REGION Network 15
   RUNG wire#powerrail
      I_Contact( "MS050-TO" )
      Coil( "MS050-TO" )
   END_RUNG
   // the same network as SCL:
   "MS050-TO" := NOT "MS050-TO";
END_REGION

REGION Network 16
   RUNG wire#powerrail
      I_Contact( "MS051-TO" )
      Coil( "MS051-TO" )
   END_RUNG
   // the same network as SCL:
   "MS051-TO" := NOT "MS051-TO";
END_REGION

REGION Network 17
   RUNG wire#powerrail
      I_Contact( "MS052-TO" )
      Coil( "MS052-TO" )
   END_RUNG
   // the same network as SCL:
   "MS052-TO" := NOT "MS052-TO";
END_REGION

REGION Network 18
   RUNG wire#powerrail
      I_Contact( "MS053-TO" )
      Coil( "MS053-TO" )
   END_RUNG
   // the same network as SCL:
   "MS053-TO" := NOT "MS053-TO";
END_REGION

REGION Network 19: Control de Iluminación Cavaleto
   RUNG wire#powerrail
      "IluminaciónMTA"()
   END_RUNG
   // the same network as SCL:
   "IluminaciónMTA"();
END_REGION
END_FUNCTION

FUNCTION "And-Byte MTA" : Void   // FC22, LAD
{ S7_Optimized_Access := 'FALSE' }
VERSION : 0.1
BEGIN

REGION Network 1
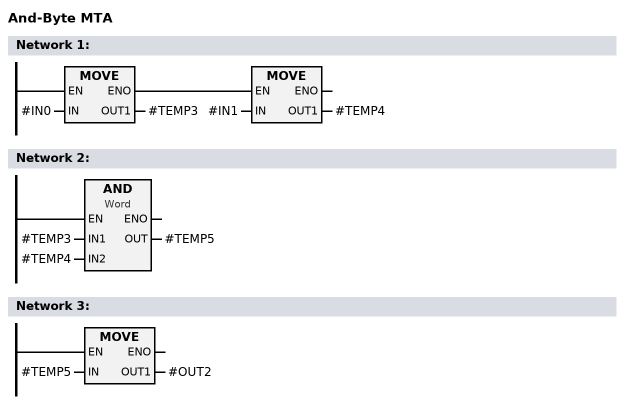
   RUNG wire#powerrail
      { S7_GenerateENO := "TRUE" } Move(in := #IN0, out1 => #TEMP3)
      { S7_GenerateENO := "TRUE" } Move(in := #IN1, out1 => #TEMP4)
   END_RUNG
   // the same network as SCL:
   // ENO of a box is taken as its EN; it also drops when the box reports an error
   #TEMP3 := #IN0;
   #TEMP4 := #IN1;
END_REGION

REGION Network 2
   RUNG wire#powerrail
      { S7_Templates := "SrcType := Word"; S7_GenerateENO := "TRUE" } And(in1 := #TEMP3, in2 := #TEMP4, out => #TEMP5)
   END_RUNG
   // the same network as SCL:
   #TEMP5 := #TEMP3 AND #TEMP4;
END_REGION

REGION Network 3
   RUNG wire#powerrail
      { S7_GenerateENO := "TRUE" } Move(in := #TEMP5, out1 => #OUT2)
   END_RUNG
   // the same network as SCL:
   #OUT2 := #TEMP5;
END_REGION
END_FUNCTION

FUNCTION "Inicialización" : Void   // FC46, LAD
{ S7_Optimized_Access := 'FALSE' }
VERSION : 0.1
BEGIN

REGION Network 1
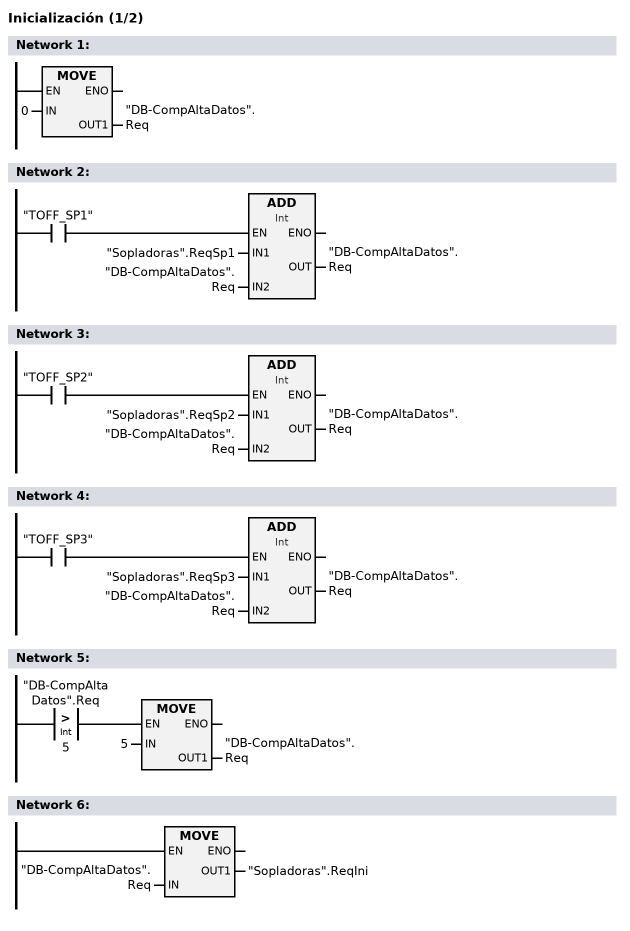
   RUNG wire#powerrail
      { S7_GenerateENO := "TRUE" } Move(in := 0, out1 => "DB-CompAltaDatos".Req)
   END_RUNG
   // the same network as SCL:
   "DB-CompAltaDatos".Req := 0;
END_REGION

REGION Network 2
   RUNG wire#powerrail
      Contact( "TOFF_SP1" )
      { S7_Templates := "SrcType := Int"; S7_GenerateENO := "TRUE" } Add(in1 := "Sopladoras".ReqSp1, in2 := "DB-CompAltaDatos".Req, out => "DB-CompAltaDatos".Req)
   END_RUNG
   // the same network as SCL:
   IF "TOFF_SP1" THEN "DB-CompAltaDatos".Req := "Sopladoras".ReqSp1 + "DB-CompAltaDatos".Req; END_IF;
END_REGION

REGION Network 3
   RUNG wire#powerrail
      Contact( "TOFF_SP2" )
      { S7_Templates := "SrcType := Int"; S7_GenerateENO := "TRUE" } Add(in1 := "Sopladoras".ReqSp2, in2 := "DB-CompAltaDatos".Req, out => "DB-CompAltaDatos".Req)
   END_RUNG
   // the same network as SCL:
   IF "TOFF_SP2" THEN "DB-CompAltaDatos".Req := "Sopladoras".ReqSp2 + "DB-CompAltaDatos".Req; END_IF;
END_REGION

REGION Network 4
   RUNG wire#powerrail
      Contact( "TOFF_SP3" )
      { S7_Templates := "SrcType := Int"; S7_GenerateENO := "TRUE" } Add(in1 := "Sopladoras".ReqSp3, in2 := "DB-CompAltaDatos".Req, out => "DB-CompAltaDatos".Req)
   END_RUNG
   // the same network as SCL:
   IF "TOFF_SP3" THEN "DB-CompAltaDatos".Req := "Sopladoras".ReqSp3 + "DB-CompAltaDatos".Req; END_IF;
END_REGION

REGION Network 5
   RUNG wire#powerrail
      { S7_Templates := "SrcType := Int" } GT_Contact(in1 := "DB-CompAltaDatos".Req, in2 := 5)
      { S7_GenerateENO := "TRUE" } Move(in := 5, out1 => "DB-CompAltaDatos".Req)
   END_RUNG
   // the same network as SCL:
   IF "DB-CompAltaDatos".Req > 5 THEN "DB-CompAltaDatos".Req := 5; END_IF;
END_REGION

REGION Network 6
   RUNG wire#powerrail
      { S7_GenerateENO := "TRUE" } Move(in := "DB-CompAltaDatos".Req, out1 => "Sopladoras".ReqIni)
   END_RUNG
   // the same network as SCL:
   "Sopladoras".ReqIni := "DB-CompAltaDatos".Req;
END_REGION

REGION Network 7
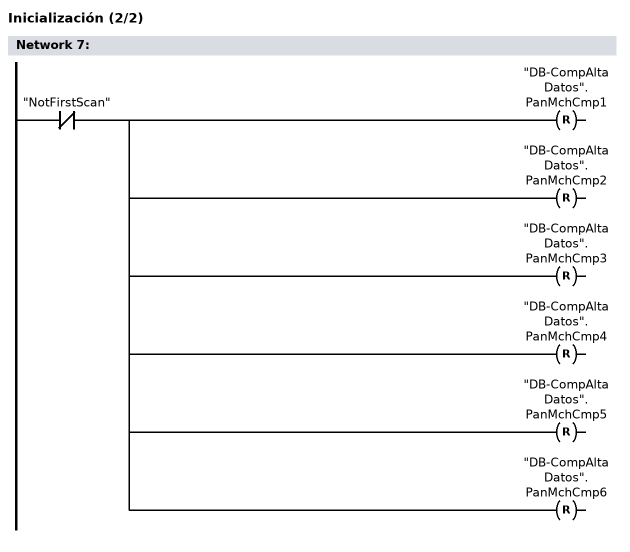
   RUNG wire#powerrail
      I_Contact( "NotFirstScan" )
      wire#w1
      R_Coil( "DB-CompAltaDatos".PanMchCmp1 )
   END_RUNG
   RUNG wire#w1
      R_Coil( "DB-CompAltaDatos".PanMchCmp2 )
   END_RUNG
   RUNG wire#w1
      R_Coil( "DB-CompAltaDatos".PanMchCmp3 )
   END_RUNG
   RUNG wire#w1
      R_Coil( "DB-CompAltaDatos".PanMchCmp4 )
   END_RUNG
   RUNG wire#w1
      R_Coil( "DB-CompAltaDatos".PanMchCmp5 )
   END_RUNG
   RUNG wire#w1
      R_Coil( "DB-CompAltaDatos".PanMchCmp6 )
   END_RUNG
   // the same network as SCL:
   IF NOT "NotFirstScan" THEN
       "DB-CompAltaDatos".PanMchCmp1 := FALSE;
       "DB-CompAltaDatos".PanMchCmp2 := FALSE;
       "DB-CompAltaDatos".PanMchCmp3 := FALSE;
       "DB-CompAltaDatos".PanMchCmp4 := FALSE;
       "DB-CompAltaDatos".PanMchCmp5 := FALSE;
       "DB-CompAltaDatos".PanMchCmp6 := FALSE;
   END_IF;
END_REGION
END_FUNCTION

// folder: Bloques Estándar

FUNCTION_BLOCK "ControladorMotoresMTA"   // FB2, LAD
{ S7_Optimized_Access := 'FALSE' }
VERSION : 0.1
BEGIN

REGION Network 2
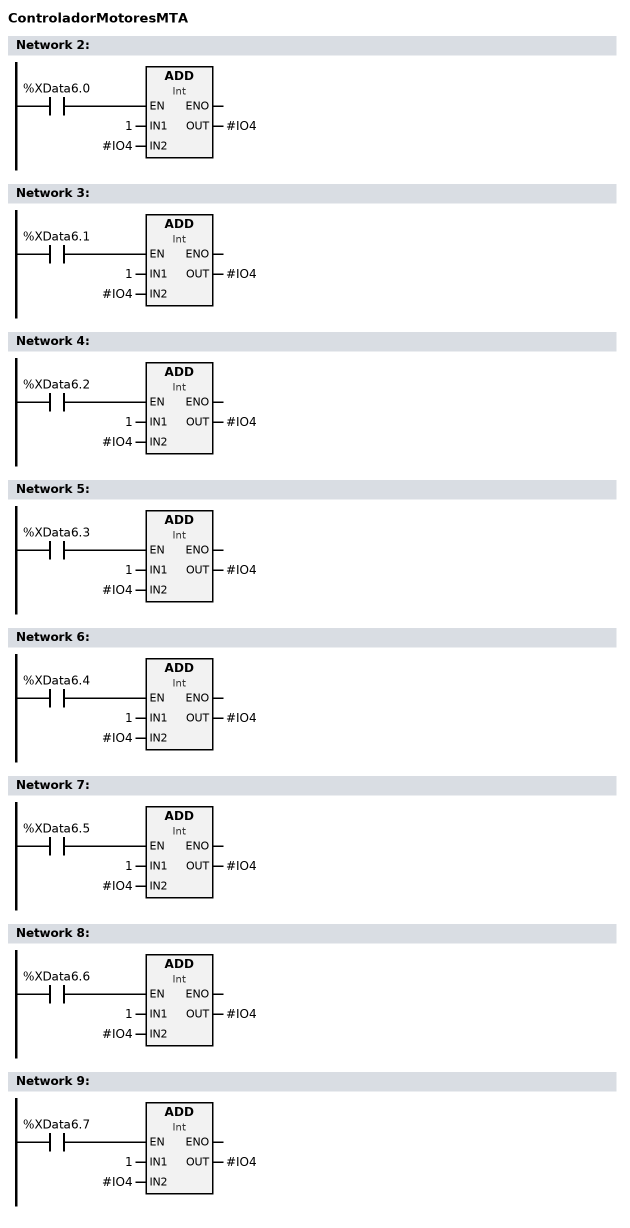
   RUNG wire#powerrail
      Contact( %XData6.0 )
      { S7_Templates := "SrcType := Int"; S7_GenerateENO := "TRUE" } Add(in1 := 1, in2 := #IO4, out => #IO4)
   END_RUNG
   // the same network as SCL:
   IF %XData6.0 THEN #IO4 := 1 + #IO4; END_IF;
END_REGION

REGION Network 3
   RUNG wire#powerrail
      Contact( %XData6.1 )
      { S7_Templates := "SrcType := Int"; S7_GenerateENO := "TRUE" } Add(in1 := 1, in2 := #IO4, out => #IO4)
   END_RUNG
   // the same network as SCL:
   IF %XData6.1 THEN #IO4 := 1 + #IO4; END_IF;
END_REGION

REGION Network 4
   RUNG wire#powerrail
      Contact( %XData6.2 )
      { S7_Templates := "SrcType := Int"; S7_GenerateENO := "TRUE" } Add(in1 := 1, in2 := #IO4, out => #IO4)
   END_RUNG
   // the same network as SCL:
   IF %XData6.2 THEN #IO4 := 1 + #IO4; END_IF;
END_REGION

REGION Network 5
   RUNG wire#powerrail
      Contact( %XData6.3 )
      { S7_Templates := "SrcType := Int"; S7_GenerateENO := "TRUE" } Add(in1 := 1, in2 := #IO4, out => #IO4)
   END_RUNG
   // the same network as SCL:
   IF %XData6.3 THEN #IO4 := 1 + #IO4; END_IF;
END_REGION

REGION Network 6
   RUNG wire#powerrail
      Contact( %XData6.4 )
      { S7_Templates := "SrcType := Int"; S7_GenerateENO := "TRUE" } Add(in1 := 1, in2 := #IO4, out => #IO4)
   END_RUNG
   // the same network as SCL:
   IF %XData6.4 THEN #IO4 := 1 + #IO4; END_IF;
END_REGION

REGION Network 7
   RUNG wire#powerrail
      Contact( %XData6.5 )
      { S7_Templates := "SrcType := Int"; S7_GenerateENO := "TRUE" } Add(in1 := 1, in2 := #IO4, out => #IO4)
   END_RUNG
   // the same network as SCL:
   IF %XData6.5 THEN #IO4 := 1 + #IO4; END_IF;
END_REGION

REGION Network 8
   RUNG wire#powerrail
      Contact( %XData6.6 )
      { S7_Templates := "SrcType := Int"; S7_GenerateENO := "TRUE" } Add(in1 := 1, in2 := #IO4, out => #IO4)
   END_RUNG
   // the same network as SCL:
   IF %XData6.6 THEN #IO4 := 1 + #IO4; END_IF;
END_REGION

REGION Network 9
   RUNG wire#powerrail
      Contact( %XData6.7 )
      { S7_Templates := "SrcType := Int"; S7_GenerateENO := "TRUE" } Add(in1 := 1, in2 := #IO4, out => #IO4)
   END_RUNG
   // the same network as SCL:
   IF %XData6.7 THEN #IO4 := 1 + #IO4; END_IF;
END_REGION
END_FUNCTION_BLOCK

// folder: Bloques Estándar/Boosters

FUNCTION "Booster (MTA)" : Void   // FC25, LAD
TITLE = Manejo General de los Boosters
{ S7_Optimized_Access := 'FALSE' }
VERSION : 0.1
   VAR_TEMP   // added for the SCL form of the ladder/FBD networks
      _w1 : Bool;
      _s5time1 : S5Time;
      _w2 : Bool;
      _s5time2 : S5Time;
      _w3 : Bool;
   END_VAR
BEGIN

REGION Network 1: Validación Horas para invertir prioridades
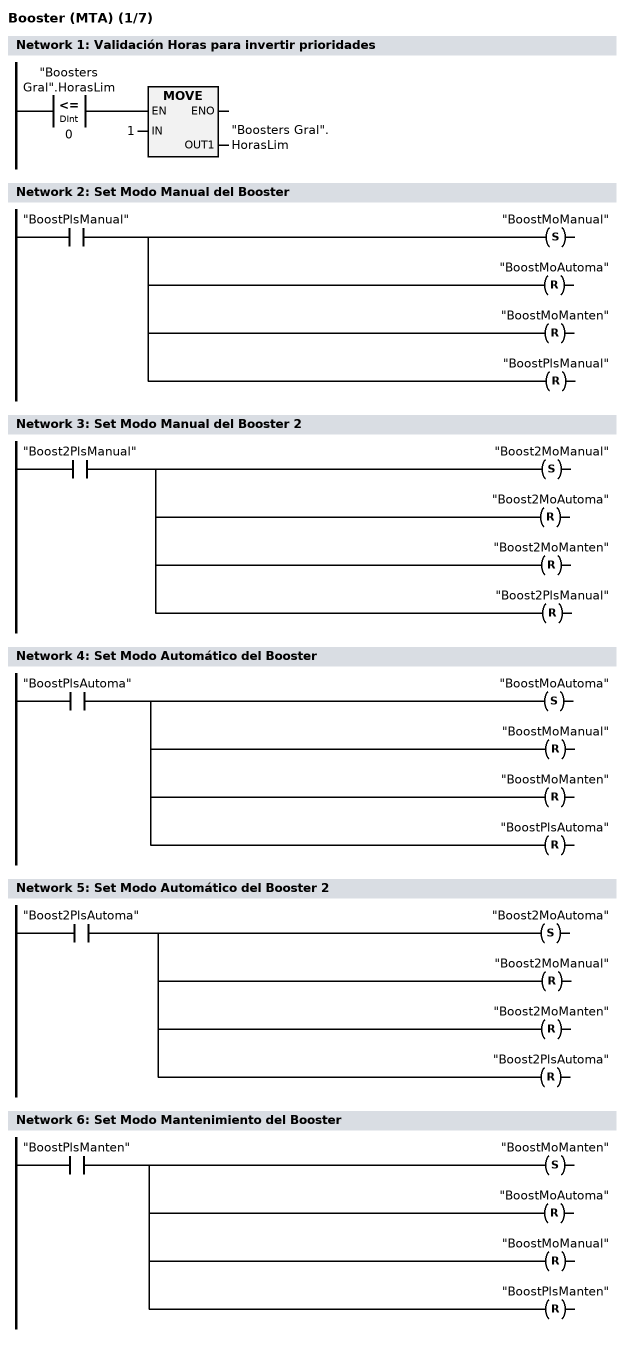
   RUNG wire#powerrail
      { S7_Templates := "SrcType := DInt" } LE_Contact(in1 := "Boosters Gral".HorasLim, in2 := 0)
      { S7_GenerateENO := "TRUE" } Move(in := 1, out1 => "Boosters Gral".HorasLim)
   END_RUNG
   // the same network as SCL:
   IF "Boosters Gral".HorasLim <= 0 THEN "Boosters Gral".HorasLim := 1; END_IF;
END_REGION

REGION Network 2: Set Modo Manual del Booster
   RUNG wire#powerrail
      Contact( "BoostPlsManual" )
      wire#w1
      S_Coil( "BoostMoManual" )
   END_RUNG
   RUNG wire#w1
      R_Coil( "BoostMoAutoma" )
   END_RUNG
   RUNG wire#w1
      R_Coil( "BoostMoManten" )
   END_RUNG
   RUNG wire#w1
      R_Coil( "BoostPlsManual" )
   END_RUNG
   // the same network as SCL:
   IF "BoostPlsManual" THEN
       "BoostMoManual" := TRUE;
       "BoostMoAutoma" := FALSE;
       "BoostMoManten" := FALSE;
       "BoostPlsManual" := FALSE;
   END_IF;
END_REGION

REGION Network 3: Set Modo Manual del Booster 2
   RUNG wire#powerrail
      Contact( "Boost2PlsManual" )
      wire#w1
      S_Coil( "Boost2MoManual" )
   END_RUNG
   RUNG wire#w1
      R_Coil( "Boost2MoAutoma" )
   END_RUNG
   RUNG wire#w1
      R_Coil( "Boost2MoManten" )
   END_RUNG
   RUNG wire#w1
      R_Coil( "Boost2PlsManual" )
   END_RUNG
   // the same network as SCL:
   IF "Boost2PlsManual" THEN
       "Boost2MoManual" := TRUE;
       "Boost2MoAutoma" := FALSE;
       "Boost2MoManten" := FALSE;
       "Boost2PlsManual" := FALSE;
   END_IF;
END_REGION

REGION Network 4: Set Modo Automático del Booster
   RUNG wire#powerrail
      Contact( "BoostPlsAutoma" )
      wire#w1
      S_Coil( "BoostMoAutoma" )
   END_RUNG
   RUNG wire#w1
      R_Coil( "BoostMoManual" )
   END_RUNG
   RUNG wire#w1
      R_Coil( "BoostMoManten" )
   END_RUNG
   RUNG wire#w1
      R_Coil( "BoostPlsAutoma" )
   END_RUNG
   // the same network as SCL:
   IF "BoostPlsAutoma" THEN
       "BoostMoAutoma" := TRUE;
       "BoostMoManual" := FALSE;
       "BoostMoManten" := FALSE;
       "BoostPlsAutoma" := FALSE;
   END_IF;
END_REGION

REGION Network 5: Set Modo Automático del Booster 2
   RUNG wire#powerrail
      Contact( "Boost2PlsAutoma" )
      wire#w1
      S_Coil( "Boost2MoAutoma" )
   END_RUNG
   RUNG wire#w1
      R_Coil( "Boost2MoManual" )
   END_RUNG
   RUNG wire#w1
      R_Coil( "Boost2MoManten" )
   END_RUNG
   RUNG wire#w1
      R_Coil( "Boost2PlsAutoma" )
   END_RUNG
   // the same network as SCL:
   IF "Boost2PlsAutoma" THEN
       "Boost2MoAutoma" := TRUE;
       "Boost2MoManual" := FALSE;
       "Boost2MoManten" := FALSE;
       "Boost2PlsAutoma" := FALSE;
   END_IF;
END_REGION

REGION Network 6: Set Modo Mantenimiento del Booster
   RUNG wire#powerrail
      Contact( "BoostPlsManten" )
      wire#w1
      S_Coil( "BoostMoManten" )
   END_RUNG
   RUNG wire#w1
      R_Coil( "BoostMoAutoma" )
   END_RUNG
   RUNG wire#w1
      R_Coil( "BoostMoManual" )
   END_RUNG
   RUNG wire#w1
      R_Coil( "BoostPlsManten" )
   END_RUNG
   // the same network as SCL:
   IF "BoostPlsManten" THEN
       "BoostMoManten" := TRUE;
       "BoostMoAutoma" := FALSE;
       "BoostMoManual" := FALSE;
       "BoostPlsManten" := FALSE;
   END_IF;
END_REGION

REGION Network 7: Set Modo Mantenimiento del Booster 2
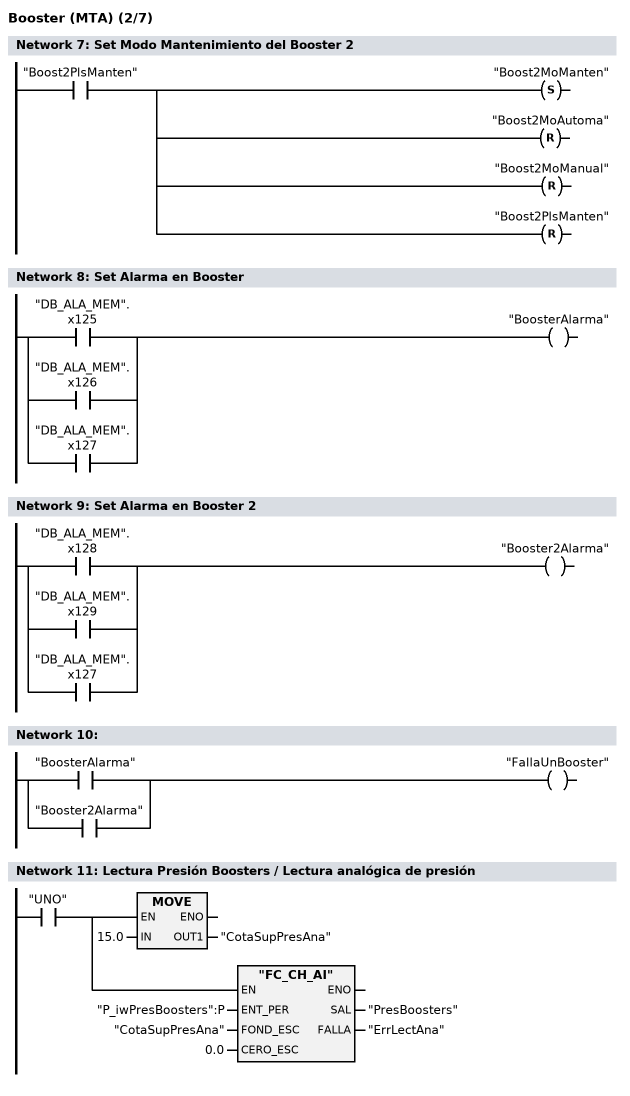
   RUNG wire#powerrail
      Contact( "Boost2PlsManten" )
      wire#w1
      S_Coil( "Boost2MoManten" )
   END_RUNG
   RUNG wire#w1
      R_Coil( "Boost2MoAutoma" )
   END_RUNG
   RUNG wire#w1
      R_Coil( "Boost2MoManual" )
   END_RUNG
   RUNG wire#w1
      R_Coil( "Boost2PlsManten" )
   END_RUNG
   // the same network as SCL:
   IF "Boost2PlsManten" THEN
       "Boost2MoManten" := TRUE;
       "Boost2MoAutoma" := FALSE;
       "Boost2MoManual" := FALSE;
       "Boost2PlsManten" := FALSE;
   END_IF;
END_REGION

REGION Network 8: Set Alarma en Booster
   RUNG wire#powerrail
      Contact( "DB_ALA_MEM".x125 )
      wire#w1
      Coil( "BoosterAlarma" )
   END_RUNG
   RUNG wire#powerrail
      Contact( "DB_ALA_MEM".x126 )
   END_RUNG wire#w1
   RUNG wire#powerrail
      Contact( "DB_ALA_MEM".x127 )
   END_RUNG wire#w1
   // the same network as SCL:
   "BoosterAlarma" := "DB_ALA_MEM".x125 OR "DB_ALA_MEM".x126 OR "DB_ALA_MEM".x127;
END_REGION

REGION Network 9: Set Alarma en Booster 2
   RUNG wire#powerrail
      Contact( "DB_ALA_MEM".x128 )
      wire#w1
      Coil( "Booster2Alarma" )
   END_RUNG
   RUNG wire#powerrail
      Contact( "DB_ALA_MEM".x129 )
   END_RUNG wire#w1
   RUNG wire#powerrail
      Contact( "DB_ALA_MEM".x127 )
   END_RUNG wire#w1
   // the same network as SCL:
   "Booster2Alarma" := "DB_ALA_MEM".x128 OR "DB_ALA_MEM".x129 OR "DB_ALA_MEM".x127;
END_REGION

REGION Network 10
   RUNG wire#powerrail
      Contact( "BoosterAlarma" )
      wire#w1
      Coil( "FallaUnBooster" )
   END_RUNG
   RUNG wire#powerrail
      Contact( "Booster2Alarma" )
   END_RUNG wire#w1
   // the same network as SCL:
   "FallaUnBooster" := "BoosterAlarma" OR "Booster2Alarma";
END_REGION

REGION Network 11: Lectura Presión Boosters / Lectura analógica de presión
   RUNG wire#powerrail
      Contact( "UNO" )
      wire#w1
      { S7_GenerateENO := "TRUE" } Move(in := 15.0, out1 => "CotaSupPresAna")
   END_RUNG
   RUNG wire#w1
      "FC_CH_AI"(ENT_PER := "P_iwPresBoosters":P, FOND_ESC := "CotaSupPresAna", CERO_ESC := 0.0, SAL => "PresBoosters", FALLA => "ErrLectAna")
   END_RUNG
   // the same network as SCL:
   IF "UNO" THEN
       "CotaSupPresAna" := 15.0;
       "FC_CH_AI"(ENT_PER := "P_iwPresBoosters":P,
                  FOND_ESC := "CotaSupPresAna",
                  CERO_ESC := 0.0,
                  SAL => "PresBoosters",
                  FALLA => "ErrLectAna");
   END_IF;
END_REGION

REGION Network 12: Bandas de presión para arranque de Boosters / Set-Reset para control analógico
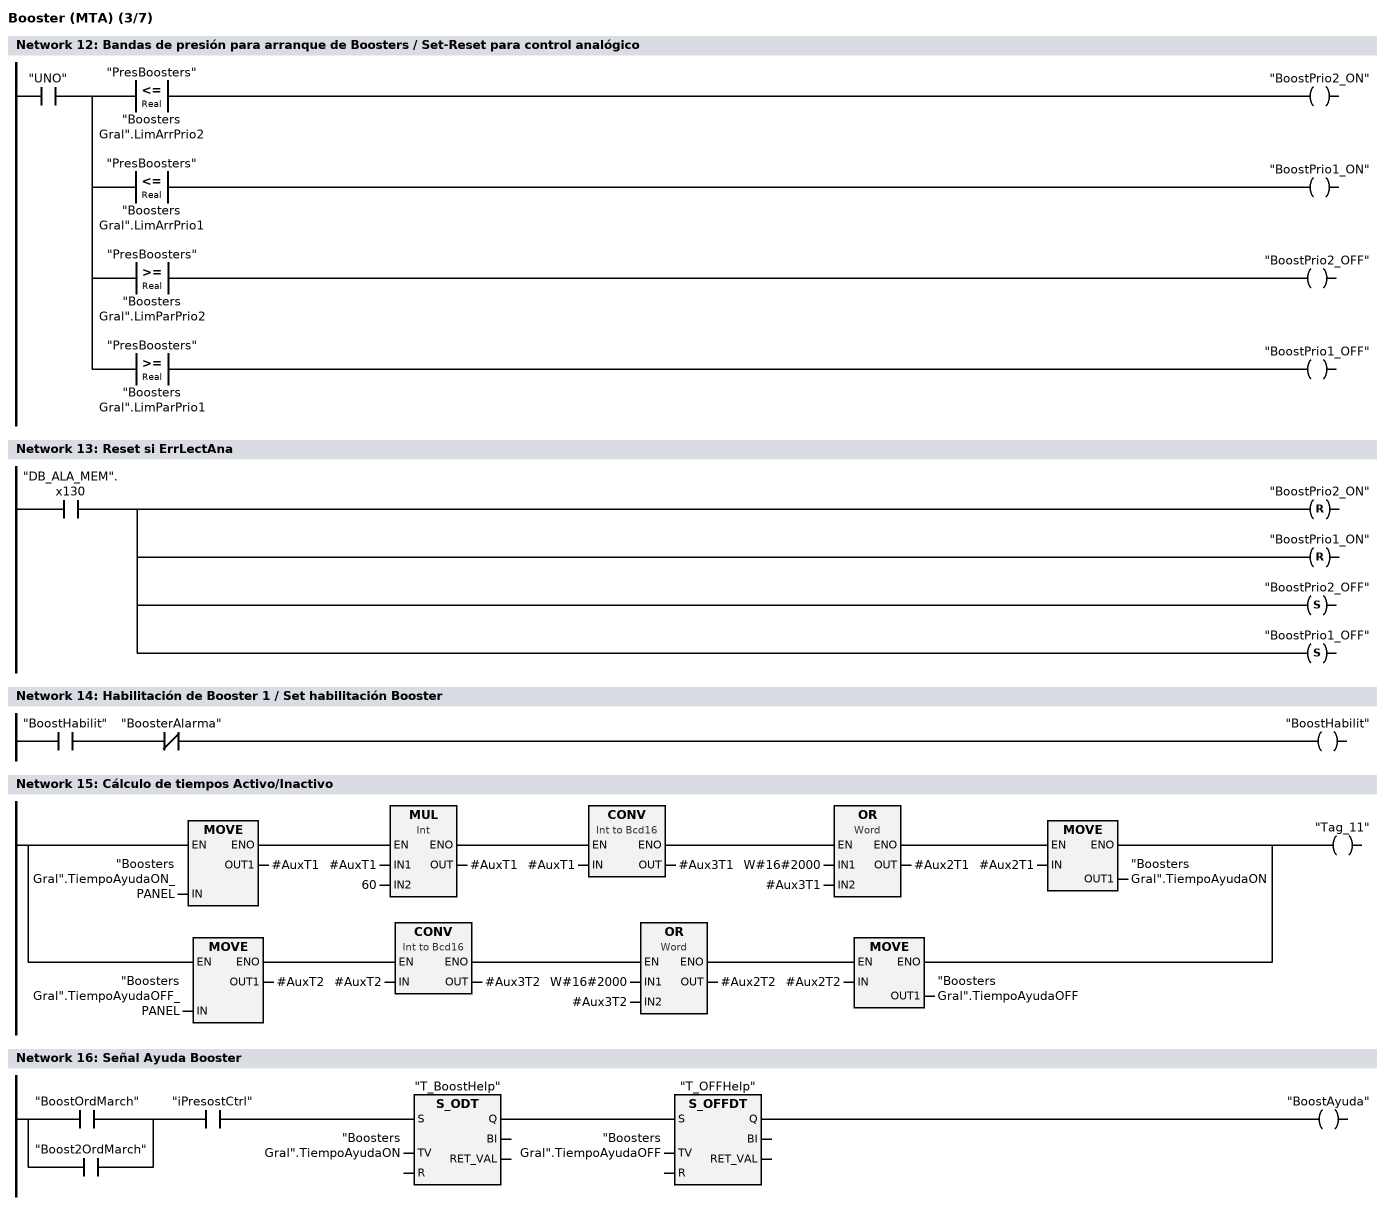
   RUNG wire#powerrail
      Contact( "UNO" )
      wire#w1
      { S7_Templates := "SrcType := Real" } LE_Contact(in1 := "PresBoosters", in2 := "Boosters Gral".LimArrPrio2)
      Coil( "BoostPrio2_ON" )
   END_RUNG
   RUNG wire#w1
      { S7_Templates := "SrcType := Real" } LE_Contact(in1 := "PresBoosters", in2 := "Boosters Gral".LimArrPrio1)
      Coil( "BoostPrio1_ON" )
   END_RUNG
   RUNG wire#w1
      { S7_Templates := "SrcType := Real" } GE_Contact(in1 := "PresBoosters", in2 := "Boosters Gral".LimParPrio2)
      Coil( "BoostPrio2_OFF" )
   END_RUNG
   RUNG wire#w1
      { S7_Templates := "SrcType := Real" } GE_Contact(in1 := "PresBoosters", in2 := "Boosters Gral".LimParPrio1)
      Coil( "BoostPrio1_OFF" )
   END_RUNG
   // the same network as SCL:
   "BoostPrio2_ON" := "UNO" AND ("PresBoosters" <= "Boosters Gral".LimArrPrio2);
   "BoostPrio1_ON" := "UNO" AND ("PresBoosters" <= "Boosters Gral".LimArrPrio1);
   "BoostPrio2_OFF" := "UNO" AND ("PresBoosters" >= "Boosters Gral".LimParPrio2);
   "BoostPrio1_OFF" := "UNO" AND ("PresBoosters" >= "Boosters Gral".LimParPrio1);
END_REGION

REGION Network 13: Reset si ErrLectAna
   RUNG wire#powerrail
      Contact( "DB_ALA_MEM".x130 )
      wire#w1
      R_Coil( "BoostPrio2_ON" )
   END_RUNG
   RUNG wire#w1
      R_Coil( "BoostPrio1_ON" )
   END_RUNG
   RUNG wire#w1
      S_Coil( "BoostPrio2_OFF" )
   END_RUNG
   RUNG wire#w1
      S_Coil( "BoostPrio1_OFF" )
   END_RUNG
   // the same network as SCL:
   IF "DB_ALA_MEM".x130 THEN
       "BoostPrio2_ON" := FALSE;
       "BoostPrio1_ON" := FALSE;
       "BoostPrio2_OFF" := TRUE;
       "BoostPrio1_OFF" := TRUE;
   END_IF;
END_REGION

REGION Network 14: Habilitación de Booster 1 / Set habilitación Booster
   RUNG wire#powerrail
      Contact( "BoostHabilit" )
      I_Contact( "BoosterAlarma" )
      Coil( "BoostHabilit" )
   END_RUNG
   // the same network as SCL:
   "BoostHabilit" := "BoostHabilit" AND NOT "BoosterAlarma";
END_REGION

REGION Network 15: Cálculo de tiempos Activo/Inactivo
   // no checked SCL form for this network; see the picture
END_REGION

REGION Network 16: Señal Ayuda Booster
   RUNG wire#powerrail
      Contact( "BoostOrdMarch" )
      wire#w1
      Contact( "iPresostCtrl" )
      S_ODT(T_NO := "T_BoostHelp", TV := "Boosters Gral".TiempoAyudaON, R :=, BI =>, RET_VAL =>)
      S_OFFDT(T_NO := "T_OFFHelp", TV := "Boosters Gral".TiempoAyudaOFF, R :=, BI =>, RET_VAL =>)
      Coil( "BoostAyuda" )
   END_RUNG
   RUNG wire#powerrail
      Contact( "Boost2OrdMarch" )
   END_RUNG wire#w1
   // the same network as SCL:
   #_s5time1 := S_ODT(T_NO := "T_BoostHelp",
                      S := ("BoostOrdMarch" OR "Boost2OrdMarch") AND "iPresostCtrl",
                      TV := "Boosters Gral".TiempoAyudaON,
                      Q => #_w1);
   #_s5time2 := S_OFFDT(T_NO := "T_OFFHelp", S := #_w1, TV := "Boosters Gral".TiempoAyudaOFF, Q => #_w2);
   "BoostAyuda" := #_w2;
END_REGION

REGION Network 17: Prioridades Boosters / Prioridades Nulas
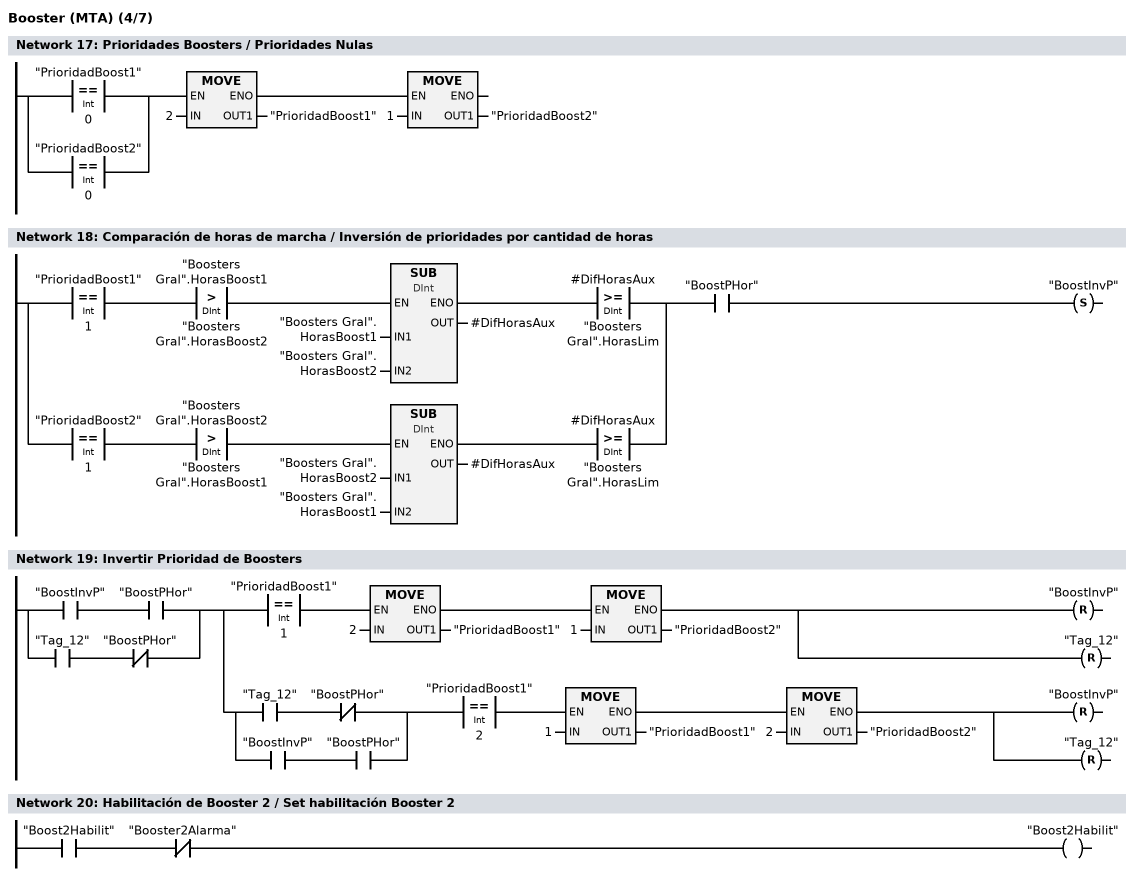
   RUNG wire#powerrail
      { S7_Templates := "SrcType := Int" } EQ_Contact(in1 := "PrioridadBoost1", in2 := 0)
      wire#w1
      { S7_GenerateENO := "TRUE" } Move(in := 2, out1 => "PrioridadBoost1")
      { S7_GenerateENO := "TRUE" } Move(in := 1, out1 => "PrioridadBoost2")
   END_RUNG
   RUNG wire#powerrail
      { S7_Templates := "SrcType := Int" } EQ_Contact(in1 := "PrioridadBoost2", in2 := 0)
   END_RUNG wire#w1
   // the same network as SCL:
   // ENO of a box is taken as its EN; it also drops when the box reports an error
   #_w1 := ("PrioridadBoost1" = 0) OR ("PrioridadBoost2" = 0);
   IF #_w1 THEN
       "PrioridadBoost1" := 2;
       "PrioridadBoost2" := 1;
   END_IF;
END_REGION

REGION Network 18: Comparación de horas de marcha / Inversión de prioridades por cantidad de horas
   RUNG wire#powerrail
      { S7_Templates := "SrcType := Int" } EQ_Contact(in1 := "PrioridadBoost1", in2 := 1)
      { S7_Templates := "SrcType := DInt" } GT_Contact(in1 := "Boosters Gral".HorasBoost1, in2 := "Boosters Gral".HorasBoost2)
      { S7_Templates := "SrcType := DInt"; S7_GenerateENO := "TRUE" } Sub(in1 := "Boosters Gral".HorasBoost1, in2 := "Boosters Gral".HorasBoost2, out => #DifHorasAux)
      { S7_Templates := "SrcType := DInt" } GE_Contact(in1 := #DifHorasAux, in2 := "Boosters Gral".HorasLim)
      wire#w1
      Contact( "BoostPHor" )
      S_Coil( "BoostInvP" )
   END_RUNG
   RUNG wire#powerrail
      { S7_Templates := "SrcType := Int" } EQ_Contact(in1 := "PrioridadBoost2", in2 := 1)
      { S7_Templates := "SrcType := DInt" } GT_Contact(in1 := "Boosters Gral".HorasBoost2, in2 := "Boosters Gral".HorasBoost1)
      { S7_Templates := "SrcType := DInt"; S7_GenerateENO := "TRUE" } Sub(in1 := "Boosters Gral".HorasBoost2, in2 := "Boosters Gral".HorasBoost1, out => #DifHorasAux)
      { S7_Templates := "SrcType := DInt" } GE_Contact(in1 := #DifHorasAux, in2 := "Boosters Gral".HorasLim)
   END_RUNG wire#w1
   // the same network as SCL:
   // ENO of a box is taken as its EN; it also drops when the box reports an error
   #_w1 := ("PrioridadBoost1" = 1) AND ("Boosters Gral".HorasBoost1 > "Boosters Gral".HorasBoost2);
   IF #_w1 THEN #DifHorasAux := "Boosters Gral".HorasBoost1 - "Boosters Gral".HorasBoost2; END_IF;
   #_w2 := ("PrioridadBoost2" = 1) AND ("Boosters Gral".HorasBoost2 > "Boosters Gral".HorasBoost1);
   #_w3 := #_w1 AND (#DifHorasAux >= "Boosters Gral".HorasLim);
   IF #_w2 THEN #DifHorasAux := "Boosters Gral".HorasBoost2 - "Boosters Gral".HorasBoost1; END_IF;
   IF (#_w3 OR (#_w2 AND (#DifHorasAux >= "Boosters Gral".HorasLim))) AND "BoostPHor" THEN
       "BoostInvP" := TRUE;
   END_IF;
END_REGION

REGION Network 19: Invertir Prioridad de Boosters
   RUNG wire#powerrail
      Contact( "BoostInvP" )
      Contact( "BoostPHor" )
      wire#w1
      { S7_Templates := "SrcType := Int" } EQ_Contact(in1 := "PrioridadBoost1", in2 := 1)
      { S7_GenerateENO := "TRUE" } Move(in := 2, out1 => "PrioridadBoost1")
      { S7_GenerateENO := "TRUE" } Move(in := 1, out1 => "PrioridadBoost2")
      wire#w2
      R_Coil( "BoostInvP" )
   END_RUNG
   RUNG wire#powerrail
      Contact( "Tag_12" )
      I_Contact( "BoostPHor" )
   END_RUNG wire#w1
   RUNG wire#w2
      R_Coil( "Tag_12" )
   END_RUNG
   RUNG wire#w1
      Contact( "Tag_12" )
      I_Contact( "BoostPHor" )
      wire#w3
      { S7_Templates := "SrcType := Int" } EQ_Contact(in1 := "PrioridadBoost1", in2 := 2)
      { S7_GenerateENO := "TRUE" } Move(in := 1, out1 => "PrioridadBoost1")
      { S7_GenerateENO := "TRUE" } Move(in := 2, out1 => "PrioridadBoost2")
      wire#w4
      R_Coil( "BoostInvP" )
   END_RUNG
   RUNG wire#w1
      Contact( "BoostInvP" )
      Contact( "BoostPHor" )
   END_RUNG wire#w3
   RUNG wire#w4
      R_Coil( "Tag_12" )
   END_RUNG
   // the same network as SCL:
   // ENO of a box is taken as its EN; it also drops when the box reports an error
   #_w1 := ("BoostInvP" AND "BoostPHor") OR ("Tag_12" AND NOT "BoostPHor");
   #_w2 := #_w1 AND ("PrioridadBoost1" = 1);
   IF #_w2 THEN
       "PrioridadBoost1" := 2;
       "PrioridadBoost2" := 1;
       "BoostInvP" := FALSE;
       "Tag_12" := FALSE;
   END_IF;
   #_w3 := #_w1 AND (("Tag_12" AND NOT "BoostPHor") OR ("BoostInvP" AND "BoostPHor")) AND ("PrioridadBoost1" = 2);
   IF #_w3 THEN
       "PrioridadBoost1" := 1;
       "PrioridadBoost2" := 2;
       "BoostInvP" := FALSE;
       "Tag_12" := FALSE;
   END_IF;
END_REGION

REGION Network 20: Habilitación de Booster 2 / Set habilitación Booster 2
   RUNG wire#powerrail
      Contact( "Boost2Habilit" )
      I_Contact( "Booster2Alarma" )
      Coil( "Boost2Habilit" )
   END_RUNG
   // the same network as SCL:
   "Boost2Habilit" := "Boost2Habilit" AND NOT "Booster2Alarma";
END_REGION

REGION Network 21: Orden de Marcha Booster
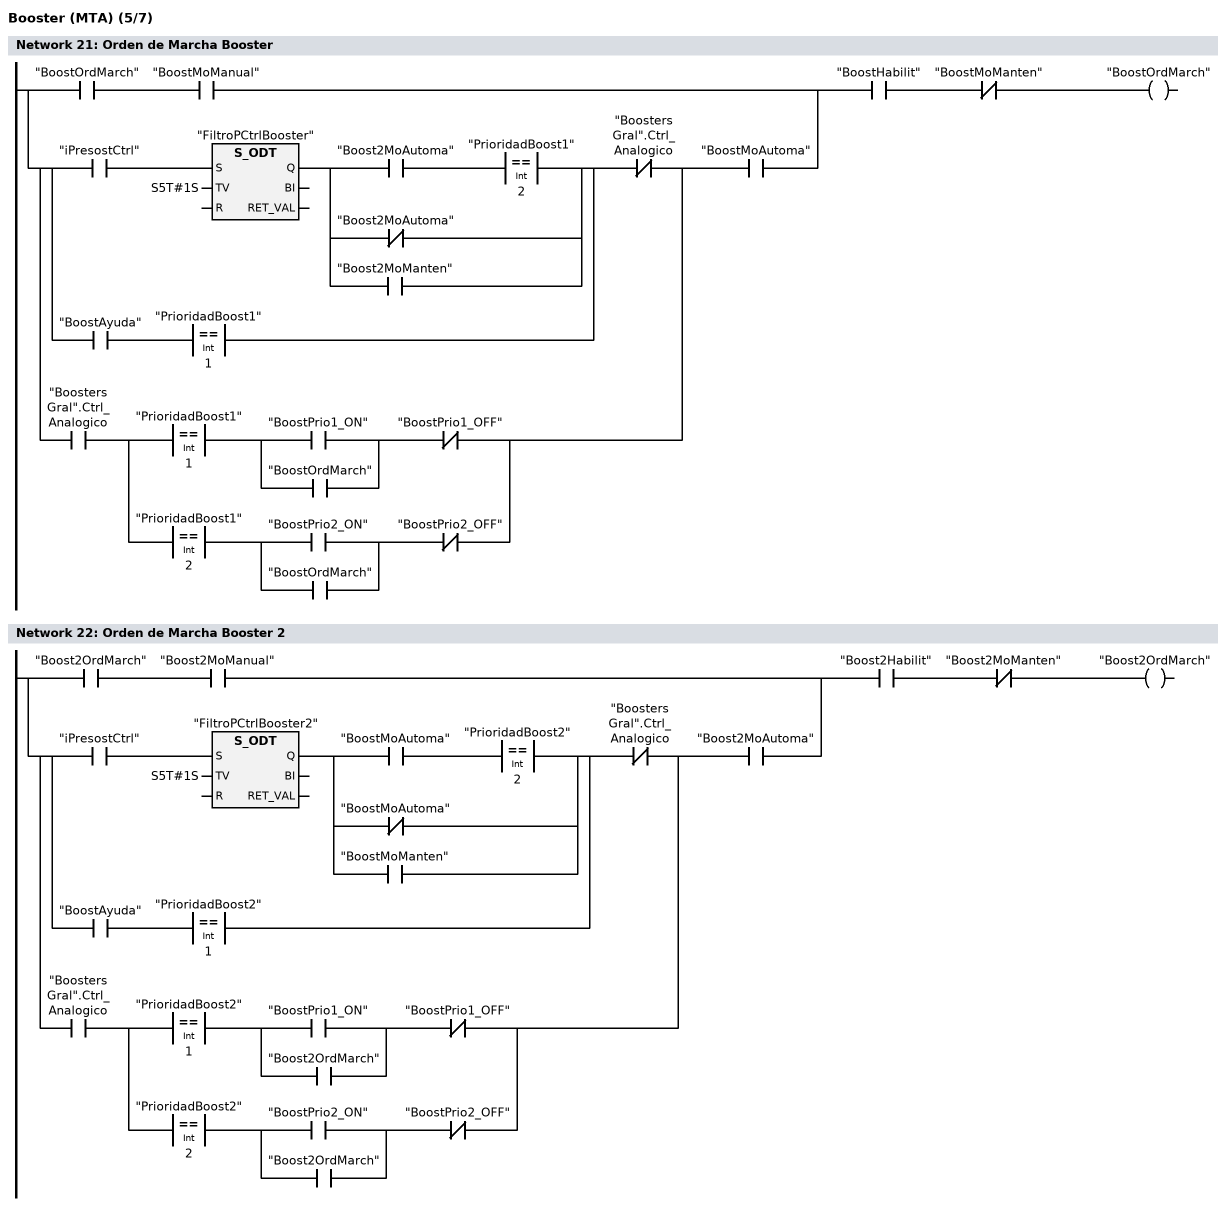
   RUNG wire#powerrail
      Contact( "BoostOrdMarch" )
      Contact( "BoostMoManual" )
      wire#w1
      Contact( "BoostHabilit" )
      I_Contact( "BoostMoManten" )
      Coil( "BoostOrdMarch" )
   END_RUNG
   RUNG wire#powerrail
      Contact( "iPresostCtrl" )
      S_ODT(T_NO := "FiltroPCtrlBooster", TV := S5T#1S, R :=, BI =>, RET_VAL =>)
      wire#w2
      Contact( "Boost2MoAutoma" )
      { S7_Templates := "SrcType := Int" } EQ_Contact(in1 := "PrioridadBoost1", in2 := 2)
      wire#w3
      I_Contact( "Boosters Gral".Ctrl_Analogico )
      wire#w4
      Contact( "BoostMoAutoma" )
   END_RUNG wire#w1
   RUNG wire#w2
      I_Contact( "Boost2MoAutoma" )
   END_RUNG wire#w3
   RUNG wire#w2
      Contact( "Boost2MoManten" )
   END_RUNG wire#w3
   RUNG wire#powerrail
      Contact( "BoostAyuda" )
      { S7_Templates := "SrcType := Int" } EQ_Contact(in1 := "PrioridadBoost1", in2 := 1)
   END_RUNG wire#w3
   RUNG wire#powerrail
      Contact( "Boosters Gral".Ctrl_Analogico )
      wire#w5
      { S7_Templates := "SrcType := Int" } EQ_Contact(in1 := "PrioridadBoost1", in2 := 1)
      wire#w6
      Contact( "BoostPrio1_ON" )
      wire#w7
      I_Contact( "BoostPrio1_OFF" )
   END_RUNG wire#w4
   RUNG wire#w6
      Contact( "BoostOrdMarch" )
   END_RUNG wire#w7
   RUNG wire#w5
      { S7_Templates := "SrcType := Int" } EQ_Contact(in1 := "PrioridadBoost1", in2 := 2)
      wire#w8
      Contact( "BoostPrio2_ON" )
      wire#w9
      I_Contact( "BoostPrio2_OFF" )
   END_RUNG wire#w4
   RUNG wire#w8
      Contact( "BoostOrdMarch" )
   END_RUNG wire#w9
   // the same network as SCL:
   #_s5time1 := S_ODT(T_NO := "FiltroPCtrlBooster", S := "iPresostCtrl", TV := S5T#1S, Q => #_w1);
   "BoostOrdMarch" := (("BoostOrdMarch" AND "BoostMoManual") OR (((((#_w1 AND (("Boost2MoAutoma" AND ("PrioridadBoost1" = 2)) OR NOT "Boost2MoAutoma" OR "Boost2MoManten")) OR ("BoostAyuda" AND ("PrioridadBoost1" = 1))) AND NOT "Boosters Gral".Ctrl_Analogico) OR ("Boosters Gral".Ctrl_Analogico AND ((("PrioridadBoost1" = 1) AND ("BoostPrio1_ON" OR "BoostOrdMarch") AND NOT "BoostPrio1_OFF") OR (("PrioridadBoost1" = 2) AND ("BoostPrio2_ON" OR "BoostOrdMarch") AND NOT "BoostPrio2_OFF")))) AND "BoostMoAutoma")) AND "BoostHabilit" AND NOT "BoostMoManten";
END_REGION

REGION Network 22: Orden de Marcha Booster 2
   RUNG wire#powerrail
      Contact( "Boost2OrdMarch" )
      Contact( "Boost2MoManual" )
      wire#w1
      Contact( "Boost2Habilit" )
      I_Contact( "Boost2MoManten" )
      Coil( "Boost2OrdMarch" )
   END_RUNG
   RUNG wire#powerrail
      Contact( "iPresostCtrl" )
      S_ODT(T_NO := "FiltroPCtrlBooster2", TV := S5T#1S, R :=, BI =>, RET_VAL =>)
      wire#w2
      Contact( "BoostMoAutoma" )
      { S7_Templates := "SrcType := Int" } EQ_Contact(in1 := "PrioridadBoost2", in2 := 2)
      wire#w3
      I_Contact( "Boosters Gral".Ctrl_Analogico )
      wire#w4
      Contact( "Boost2MoAutoma" )
   END_RUNG wire#w1
   RUNG wire#w2
      I_Contact( "BoostMoAutoma" )
   END_RUNG wire#w3
   RUNG wire#w2
      Contact( "BoostMoManten" )
   END_RUNG wire#w3
   RUNG wire#powerrail
      Contact( "BoostAyuda" )
      { S7_Templates := "SrcType := Int" } EQ_Contact(in1 := "PrioridadBoost2", in2 := 1)
   END_RUNG wire#w3
   RUNG wire#powerrail
      Contact( "Boosters Gral".Ctrl_Analogico )
      wire#w5
      { S7_Templates := "SrcType := Int" } EQ_Contact(in1 := "PrioridadBoost2", in2 := 1)
      wire#w6
      Contact( "BoostPrio1_ON" )
      wire#w7
      I_Contact( "BoostPrio1_OFF" )
   END_RUNG wire#w4
   RUNG wire#w6
      Contact( "Boost2OrdMarch" )
   END_RUNG wire#w7
   RUNG wire#w5
      { S7_Templates := "SrcType := Int" } EQ_Contact(in1 := "PrioridadBoost2", in2 := 2)
      wire#w8
      Contact( "BoostPrio2_ON" )
      wire#w9
      I_Contact( "BoostPrio2_OFF" )
   END_RUNG wire#w4
   RUNG wire#w8
      Contact( "Boost2OrdMarch" )
   END_RUNG wire#w9
   // the same network as SCL:
   #_s5time1 := S_ODT(T_NO := "FiltroPCtrlBooster2", S := "iPresostCtrl", TV := S5T#1S, Q => #_w1);
   "Boost2OrdMarch" := (("Boost2OrdMarch" AND "Boost2MoManual") OR (((((#_w1 AND (("BoostMoAutoma" AND ("PrioridadBoost2" = 2)) OR NOT "BoostMoAutoma" OR "BoostMoManten")) OR ("BoostAyuda" AND ("PrioridadBoost2" = 1))) AND NOT "Boosters Gral".Ctrl_Analogico) OR ("Boosters Gral".Ctrl_Analogico AND ((("PrioridadBoost2" = 1) AND ("BoostPrio1_ON" OR "Boost2OrdMarch") AND NOT "BoostPrio1_OFF") OR (("PrioridadBoost2" = 2) AND ("BoostPrio2_ON" OR "Boost2OrdMarch") AND NOT "BoostPrio2_OFF")))) AND "Boost2MoAutoma")) AND "Boost2Habilit" AND NOT "Boost2MoManten";
END_REGION

REGION Network 23: Motor Booster 1 / Bloque de Motor Booster
